      // Drži izdelek v vrteči mizi
              R    "Y3/3_OdpiranjeDržalaKomada"
   END_STEP
   TRANSITION Trans34 FROM ("Odpri klešče", "DRŽI IZDELEK") TO ("VRAČANJE NAZAJ", "Odmik konusa")   // T34
      := "PrijemaloKontaktaOdprto" AND "DrzanjeKontakta";
   END_TRANSITION
   STEP "VRAČANJE NAZAJ":   // S9, max time T#10S, warning time T#7S
      supervision V := (NOT "PrijemaloKontaktaOdprto" OR NOT "SDAT1".oPoz1Dosezena) AND (#"VRAČANJE NAZAJ".T > t#2000MS);
              S    "Y2/1_NalaganjeNazanj"
              R    "Y2/1_NalaganjeNaprej"
              R    "Y1/3_OdmičniCilinderKonusa"
   END_STEP
   TRANSITION Trans41 FROM ("Odmik konusa", "VRAČANJE NAZAJ") TO ("ZAVRTI MIZO", Step36)   // T41
      := ((("FB_KEYENCE_GT2_odmikKonusaKroznika".out >= 57000) AND ("FB_KEYENCE_GT2_ODMIKVARJENJA".out >= 39000)) OR ("AlwaysFALSE" AND "FB_KEYENCE_GT2_ODMIKVARJENJA".oPoz1Dosezena AND "FB_KEYENCE_GT2_odmikKonusaKroznika".oPoz1Dosezena)) AND ("FB_AKD_VrtenjeKroznika".o_BerrStatus = 1);
   END_TRANSITION
   STEP "ZAVRTI MIZO":   // S10, max time T#10S, warning time T#7S
      interlock C := "PozKontaktNazaj" AND "DrzanjeIzmetKontakta" AND "IzmetKontaktaNazaj" AND "PozKontaktNazaj" AND "Y1/4_odmičniCilinderVarjenje_GOR";
      (C)     S    "db_AKD".KROZNIK.PODATKI.ServoGo
   END_STEP
   STEP "ZAKLEP KONUSA":   // S11, max time T#10S, warning time T#7S
              S    "Y1/3_OdmičniCilinderKonusa"
   END_STEP
   STEP "PODAJANJE PLOŠČICE":   // S14, max time T#10S, warning time T#7S
      supervision V := (NOT "SDAT1".oPoz1Dosezena OR NOT "PozKontaktNaKoncuLetve") AND (#"PODAJANJE PLOŠČICE".T > t#2000MS);
              S    "Y2/1_dovajanjePlosciceNazaj"
              R    "Y2_1_dovajanjePlosciceNaprej"
   END_STEP
   TRANSITION Trans38 FROM "PODAJANJE PLOŠČICE" TO "ZAČETEK NOVEGA CIKLA"   // T38: SDAT VREDNOSTI <> 0
      := "SDAT1".oPoz1Dosezena AND "PozKontaktNaKoncuLetve" AND ("SDAT1".out <> 0.0) AND ("SDAT2".out <> 0.0);
   END_TRANSITION
   STEP Step36:   // S36, max time T#10S, warning time T#7S
      interlock C := "PozKontaktNaKoncuLetve" AND "SDAT1".oPoz1Dosezena;
      // Zapri prijemalo
      (C)     R    "Y3/1_PrijemaloKontaktaOdpri"
   END_STEP
   TRANSITION Trans43 FROM ("ZAVRTI MIZO", Step36) TO (Step40, Step37)   // T43
      := NOT "db_AKD".KROZNIK.PODATKI.ServoGo AND "TON_MOTOR".Q AND "DB_PODATKI".KROZNA_MIZA.IzdelekPrisotenArray[5];
   END_TRANSITION
   TRANSITION Trans55 FROM ("ZAVRTI MIZO", Step36) TO "Izdelek ni bil prisoten"   // T55
      := NOT "db_AKD".KROZNIK.PODATKI.ServoGo AND "TON_MOTOR".Q AND NOT "DB_PODATKI".KROZNA_MIZA.IzdelekPrisotenArray[5];
   END_TRANSITION
   STEP "Zakasnitev varjenja":   // S35, max time T#10S, warning time T#7S
      supervision V := ((NOT "EndOfSequency_WC" AND "AlwaysFALSE") OR NOT "FB_KEYENCE_GT2_ODMIKVARJENJA".oPoz4Dosezena) AND (#"Zakasnitev varjenja".T > t#2000MS);
   END_STEP
   TRANSITION Trans19 FROM "Zakasnitev varjenja" TO "Dvig elektrode"   // T19
      := ("EndOfSequency_WC" AND NOT "WeldFault" AND "FB_KEYENCE_GT2_ODMIKVARJENJA".oPoz4Dosezena) OR ("WeldFault" AND "FB_KEYENCE_GT2_ODMIKVARJENJA".oPoz4Dosezena) OR NOT "ExternalWeldOn";
   END_TRANSITION
   STEP "ZAČETEK NOVEGA CIKLA":   // S31, max time T#10S, warning time T#7S
      supervision V := (NOT "PozKontaktNaKoncuLetve" OR NOT "PrisotnostTraka" OR NOT "FB_IOL_IFM_SV_DB".oPretokOK OR NOT "FB_IOL_IFM_SV_DB".oTempOK OR "NapakaCiscenjaElektrode" OR "NapakaOdvijanjaTrau" OR ("FB_TekociTrak_DB".stat_skatla1Polna AND "FB_TekociTrak_DB".stat_skatla2Polna)) AND (#"ZAČETEK NOVEGA CIKLA".T > t#2000MS);
   END_STEP
   TRANSITION Trans48 FROM "ZAČETEK NOVEGA CIKLA" TO Step38   // T48
      := NOT "STEVEC_KONEC_TRAKA_DOSEZEN" AND "FB_IOL_IFM_SV_DB".oPretokOK AND "FB_IOL_IFM_SV_DB".oTempOK AND NOT "NapakaCiscenjaElektrode" AND NOT "NapakaOdvijanjaTrau" AND (NOT "FB_TekociTrak_DB".stat_skatla1Polna OR NOT "FB_TekociTrak_DB".stat_skatla2Polna);
   END_TRANSITION
   STEP Step38:   // S38, max time T#10S, warning time T#7S
      supervision V := NOT "PozKontaktNaKoncuLetve" AND (#Step38.T > t#3000MS);
   END_STEP
   TRANSITION Trans45 FROM Step38 TO Step43   // T45
      := "SDAT1".oPoz1Dosezena AND "PozKontaktNaKoncuLetve" AND NOT "DB_PODATKI".KROZNA_MIZA.IzdelekPrisoten.%X7;
   END_TRANSITION
   TRANSITION Trans47 FROM Step38 TO Step41   // T47: Izdelek prisoten v mizi
      := "DB_PODATKI".KROZNA_MIZA.IzdelekPrisoten.%X7;
   END_TRANSITION
   STEP Step43:   // S43, max time T#10S, warning time T#7S
              R    "DB_VARJENJE".PODATKI.input.ZajtevaZaVarjenje
   END_STEP
   TRANSITION Trans52 FROM Step43 TO ("Odpri Držanje komada", "Zapiranje klešč")   // T52
      := #Step43.T > t#20MS;
   END_TRANSITION
   STEP IZMET:   // S32, max time T#10S, warning time T#7S
              L    "Y4/3_OdpiranjeIzmetaKontakta",T#50mS
              L    "Y5/3_IzmetKomadov", T#50mS
   END_STEP
   TRANSITION Trans46 FROM IZMET TO "NALAGANJE PLOŠČICE/KOMADA"   // T46
      := (#IZMET.T > t#100MS) AND "SDAT1".oPoz1Dosezena;
   END_TRANSITION
   STEP Step41:   // S41, max time T#10S, warning time T#7S
   END_STEP
   TRANSITION Trans49 FROM Step41 TO ("VRAČANJE NAZAJ", "Odmik konusa")   // T49
      := #Step41.T > t#20MS;
   END_TRANSITION
   STEP Step30:   // S30, max time T#10S, warning time T#7S
   END_STEP
   TRANSITION Trans22 FROM Step30 TO "POZ ZAVARJENO"   // T22
      := TRUE;
   END_TRANSITION
   STEP Step37:   // S37, max time T#10S, warning time T#7S
   END_STEP
   TRANSITION Trans37 FROM Step37 TO ("ZAKLEP KONUSA", "IZMET KOSOV", "Poravnava Naprej_1", "Vlaganje ploščice_1", PODAJANJE_1)   // T37: Počakaj da se motor odvrti
      := (#Step37.T > t#20MS) AND ("DB_PODATKI".KROZNA_MIZA.IzdelekPrisoten.%X7 OR "AlwaysTRUE") AND "FB_AKD_DB_RezanjePodajanje".iAKD.PODATKI_TO_SIEMENS.DriveStopen;
   END_TRANSITION
   STEP Step40:   // S40, max time T#10S, warning time T#7S
      supervision V := NOT "PozKontaktNaKoncuLetve" AND (#Step40.T > t#2000MS);
   END_STEP
   TRANSITION Trans44 FROM Step40 TO ("Zapiranje klešč_1", "Odpri Držanje komada_1", "ZAKLEP KONUSA_1")   // T44
      := NOT "DB_PODATKI".KROZNA_MIZA.IzdelekPrisoten.%X7 AND (#Step40.T > t#20MS) AND "PozKontaktNaKoncuLetve";
   END_TRANSITION
   TRANSITION Trans53 FROM Step40 TO "VRAČANJE NAZAJ_1"   // T53
      := "AlwaysTRUE" AND (#Step40.T > t#100MS) AND "DB_PODATKI".KROZNA_MIZA.IzdelekPrisoten.%X7;
   END_TRANSITION
   STEP "Odpri klešče_1":   // S21, max time T#10S, warning time T#7S
      supervision V := NOT "PrijemaloKontaktaOdprto" AND (#"Odpri klešče_1".T > t#2000MS);
              S    "Y3/1_PrijemaloKontaktaOdpri"
              S    "DB_PODATKI".KROZNA_MIZA.IzdelekPrisoten.%X7
   END_STEP
   STEP "Vstavljanje v mizo_1":   // S15, max time T#10S, warning time T#7S
      interlock C := "FB_KEYENCE_GT2_odmikKonusaKroznika".oPoz2Dosezena;
      supervision V := (NOT "PrijemaloKontaktaZaprto" OR NOT "SDAT1".oPoz2Dosezena) AND (#"Vstavljanje v mizo_1".T > t#2000MS);
      (C)     S    "Y2/1_NalaganjeNaprej"
              R    "Y2/1_NalaganjeNazanj"
   END_STEP
   TRANSITION Trans35 FROM "Vstavljanje v mizo_1" TO Step42   // T35
      := "PrijemaloKontaktaZaprto" AND "SDAT1".oPoz2Dosezena;
   END_TRANSITION
   STEP "Zapiranje klešč_1":   // S6, max time T#10S, warning time T#7S
      interlock C := "PozKontaktNaKoncuLetve";
      (C)     R    "Y3/1_PrijemaloKontaktaOdpri"
   END_STEP
   STEP "Odpri Držanje komada_1":   // S13, max time T#10S, warning time T#7S
      supervision V := "DrzanjeKontakta" AND (#"Odpri Držanje komada_1".T > t#2000MS);
      // OdpriDržanjeKomada -
              S    "Y3/3_OdpiranjeDržalaKomada"
   END_STEP
   STEP "DRŽI IZDELEK_1":   // S33, max time T#10S, warning time T#7S
      supervision V := NOT "DrzanjeKontakta" AND (#"DRŽI IZDELEK_1".T > t#2000MS);
      // Drži izdelek v vrteči mizi
              R    "Y3/3_OdpiranjeDržalaKomada"
   END_STEP
   TRANSITION Trans40 FROM ("Odpri klešče_1", "DRŽI IZDELEK_1") TO "VRAČANJE NAZAJ_1"   // T40
      := "PrijemaloKontaktaOdprto" AND "DrzanjeKontakta";
   END_TRANSITION
   STEP "VRAČANJE NAZAJ_1":   // S34, max time T#10S, warning time T#7S
      supervision V := (NOT "PrijemaloKontaktaOdprto" OR NOT "SDAT1".oPoz1Dosezena) AND (#"VRAČANJE NAZAJ_1".T > t#2000MS);
              S    "Y2/1_NalaganjeNazanj"
              R    "Y2/1_NalaganjeNaprej"
   END_STEP
   STEP "ZAKLEP KONUSA_1":   // S39, max time T#10S, warning time T#7S
              S    "Y1/3_OdmičniCilinderKonusa"
   END_STEP
   TRANSITION Trans33 FROM ("Zapiranje klešč_1", "Odpri Držanje komada_1", "ZAKLEP KONUSA_1") TO "Vstavljanje v mizo_1"   // T33: Prijemalo zaprto
      := "PrijemaloKontaktaZaprto" AND NOT "DrzanjeKontakta" AND "ZaporaIzdelka";
   END_TRANSITION
   STEP Step42:   // S42, max time T#10S, warning time T#7S
              S    "Y3/1_PrijemaloKontaktaOdpri"
              S    "DB_PODATKI".KROZNA_MIZA.IzdelekPrisoten.%X7
   END_STEP
   TRANSITION Trans54 FROM Step42 TO ("DRŽI IZDELEK_1", "Odpri klešče_1")   // T54
      := TRUE;
   END_TRANSITION
   STEP "Izdelek ni bil prisoten":   // S44, max time T#10S, warning time T#7S
   END_STEP
   TRANSITION Trans56 FROM "Izdelek ni bil prisoten" TO "ZAČETEK NOVEGA CIKLA"   // T56, jump
      := TRUE;
   END_TRANSITION
   STEP "Poravnava Naprej_1":   // S46, max time T#10S, warning time T#7S
              S    "Y2/3_PozicioniranjeKontaktovNaprej"
              R    "Y2/3_PozicioniranjeKontaktovNazaj"
              S    "1Y1_OdklepZapore"
   END_STEP
   STEP "Vlaganje ploščice_1":   // S48, max time T#10S, warning time T#7S
      interlock C := "FB_KEYENCE_GT2_ODMIKVARJENJA".oPoz1Dosezena;
      supervision V := NOT "SDAT2".oPoz2Dosezena AND (#"Vlaganje ploščice_1".U > t#2000MS);
              S    "Y2_1_dovajanjePlosciceNaprej"
              R    "Y2/1_dovajanjePlosciceNazaj"
   END_STEP
   STEP "ZVAR NOK":   // S50, max time T#10S, warning time T#7S
      supervision V := "IEC_Counter_0_DB_1".QU;
              R    "DB_PODATKI".KROZNA_MIZA.IzdelekZavarjen.%X5
              N    "DB_PODATKI".KROZNA_MIZA.StatusIzdelkaVarjenje[5] := 1
              S    "DB_HMI".Varjenje.ResetWithWC
   END_STEP
   TRANSITION Trans59 FROM "ZVAR NOK" TO "Zakasnitev varjenja"   // T59
      := NOT "IEC_Counter_0_DB_1".QU;
   END_TRANSITION
   STEP "Zvar  OK":   // S51, max time T#10S, warning time T#7S
              S    "DB_PODATKI".KROZNA_MIZA.IzdelekZavarjen.%X5
              N    "DB_PODATKI".KROZNA_MIZA.StatusIzdelkaVarjenje[5] := 10
   END_STEP
   TRANSITION Trans60 FROM "Zvar  OK" TO "Zakasnitev varjenja"   // T60
      := TRUE;
   END_TRANSITION
   STEP Step52:   // S52, max time T#10S, warning time T#7S
   END_STEP
   TRANSITION Trans62 FROM Step52 TO (Step45, REZANJE)   // T62
      := TRUE;
   END_TRANSITION
   STEP Step16:   // S16, max time T#10S, warning time T#7S
      supervision V := NOT "EndOfSequency_WC" AND (#Step16.T > t#1000MS);
   END_STEP
   TRANSITION Trans50 FROM Step16 TO "Zvar  OK"   // T50
      := "EndOfSequency_WC" AND NOT "WeldFault";
   END_TRANSITION
   TRANSITION Trans58 FROM Step16 TO "ZVAR NOK"   // T58
      := "WeldFault";
   END_TRANSITION
   STEP Step54:   // S54, max time T#10S, warning time T#7S
      // Ploščica Odrezana - setiraj bit
              N    "db_AKD".REZANJEPODAJANJE.PODATKI.PloscicaOdrezana := True
   END_STEP
   TRANSITION Trans64 FROM Step54 TO END   // T64
      := TRUE;
   END_TRANSITION
   STEP "RESET VSEGA":   // S2, max time T#10S, warning time T#7S
      // RESET ENOTE
              R    "Y2/1_NalaganjeNaprej"
              R    "Y2/1_NalaganjeNazanj"
              S    "Y3/1_PrijemaloKontaktaOdpri"
              R    "Y2/3_PozicioniranjeKontaktovNazaj"
              S    "Y1/3_OdmičniCilinderKonusa"
              R    "Y3/3_OdpiranjeDržalaKomada"
              R    "Y4/3_OdpiranjeIzmetaKontakta"
              R    "Y5/3_IzmetKomadov"
              S    "Y1/4_odmičniCilinderVarjenje_GOR"
              S    "1Y1_OdklepZapore"
              S    "Y2/1_dovajanjePlosciceNazaj"
              R    "Y2_1_dovajanjePlosciceNaprej"
              R    "db_AKD".REZANJEPODAJANJE.PODATKI.Odrezano
              R    "db_AKD".REZANJEPODAJANJE.PODATKI.Podano
              R    "Y2/1_dovajanjePlosciceNazaj"
              R    "Y2_1_dovajanjePlosciceNaprej"
              R    "Y2/3_PozicioniranjeKontaktovNaprej"
              S    "Y2/3_PozicioniranjeKontaktovNazaj"
              R    "Y2_1_dovajanjePlosciceNaprej"
              R    "Y2/1_dovajanjePlosciceNazaj"
              R    "db_AKD".REZANJEPODAJANJE.PODATKI.Odrezano
              R    "db_AKD".REZANJEPODAJANJE.PODATKI.Podano
              R    "db_AKD".REZANJEPODAJANJE.PODATKI.ZahtevaPoPodajanju
              R    "db_AKD".REZANJEPODAJANJE.PODATKI.ZahtevaPoRezanju
              R    "DB_VARJENJE".PODATKI.input.ZajtevaZaVarjenje
              R    "Y1/4_odmičniCilinderVarjenjeDOL"
              S    "Y3/1_PrijemaloKontaktaOdpri"
              R    "DB_VARJENJE".PODATKI.input.ZajtevaZaVarjenje
              R    "DB_HMI".Varjenje.ResetWithWC
              R    "Y5/3_IzmetKomadov"
   END_STEP
   TRANSITION Trans28 FROM "RESET VSEGA" TO IZMET   // T28: OK
      := TRUE;
   END_TRANSITION
   STEP "Odmik vilic":   // S27, max time T#10S, warning time T#7S
      supervision V := (NOT "SDAT2".oPoz1Dosezena OR (NOT "TimerReady" AND "AlwaysFALSE") OR ("WeldFault" AND "AlwaysFALSE") OR NOT "SpotSelectionTakeOver") AND (#"Odmik vilic".T > t#2000MS);
              S    "Y2/1_dovajanjePlosciceNazaj"
              R    "Y2_1_dovajanjePlosciceNaprej"
              N    "db_AKD".REZANJEPODAJANJE.PODATKI.PloscicaOdrezana := false
   END_STEP
   TRANSITION Trans26 FROM ("VRAČANJE NAZAJ_1", "Poravnava nazaj", "Odmik vilic") TO (Varjenje, Step52)   // T26: Vilice v izhodišču + pdoajanje v izhodišču
      := ("SDAT2".oPoz1Dosezena OR ("SDAT2".out <= 60.0)) AND "PozKontaktNazaj" AND (("TimerReady" AND NOT "WeldFault") OR "AlwaysTRUE") AND "SpotSelectionTakeOver" AND "FB_KEYENCE_GT2_ODMIKVARJENJA".oPoz3Dosezena AND ("SDAT1".oPoz1Dosezena OR ("SDAT1".out <= 50.0) OR "AlwaysTRUE") AND "FB_KEYENCE_GT2_odmikKonusaKroznika".oPoz2Dosezena AND ("FB_AKD_DB_RezanjePodajanje".o_BerrStatus = 1);
   END_TRANSITION
   STEP "Odmik konusa":   // S22, max time T#10S, warning time T#7S
              R    "Y1/3_OdmičniCilinderKonusa"
   END_STEP
   STEP PODAJANJE_1:   // S47, max time T#10S, warning time T#7S
              S    "db_AKD".REZANJEPODAJANJE.PODATKI.Podano
              L    "db_AKD".REZANJEPODAJANJE.PODATKI.ZahtevaPoPodajanju, T#50mS
   END_STEP
   TRANSITION Trans36 FROM PODAJANJE_1 TO Step53   // T36
      := NOT "FB_AKD_DB_RezanjePodajanje".bServoGo AND "TON_REZANJEPODAJANJE".Q AND NOT "db_AKD".REZANJEPODAJANJE.PODATKI.vPODAJANJU AND (#PODAJANJE_1.T > t#10MS);
   END_TRANSITION
   STEP Step53:   // S53, max time T#10S, warning time T#7S
   END_STEP
   TRANSITION Trans24 FROM ("IZMET KOSOV", "ZAKLEP KONUSA", "Poravnava Naprej_1", "Vlaganje ploščice_1", Step53) TO "Spust Elektrode"   // T24: Izmet Nazaj in KONUS zaklenjen
      := "DrzanjeIzmetKontakta" AND "IzmetKontaktaNazaj" AND "FB_KEYENCE_GT2_odmikKonusaKroznika".oPoz2Dosezena AND "PozKontaktNaprej" AND "SDAT2".oPoz2Dosezena AND (#"IZMET KOSOV".T > t#50MS);
   END_TRANSITION
   STEP Step49:   // S49, max time T#10S, warning time T#7S
              S    "Y2_1_dovajanjePlosciceNaprej"
              R    "Y2/1_dovajanjePlosciceNazaj"
   END_STEP
   TRANSITION Trans51 FROM Step49 TO "Izdelek ni bil prisoten"   // T51
      := TRUE;
   END_TRANSITION

   // permanent post-instructions
   NETWORK 1
   TITLE = ODKLENI LIN PROGO
      "1Y1_OdklepZapore" := ("SDAT1".out >= 19.5) OR (("SDAT1".out < 19.5) AND NOT "PozKontaktNaKoncuLetve");
   NETWORK 2
   TITLE = VSTAVLJANJE KOSA V MIZO
   NETWORK 3
      IF "AlwaysFALSE" THEN
          "FB_Alarms_DB_1"(I_FAULT_RESET := "ResetNapake",   // "FB_Alarms"
                           I_Alarm_0 := "FB_GL_PROGRAM_DB"."Spust Elektrode".X AND NOT "FB_KEYENCE_GT2_ODMIKVARJENJA".bBDC3,
                           I_Alarm_1 := ("FB_FESTO_SDE1_DB".oPritisk < 6.0) AND "AlwaysFALSE",
                           I_Alarm_2 := NOT "PrisotnostTraka" AND "AlwaysFALSE",
                           I_Alarm_3 := #"Vstavljanje v mizo_1".VA,
                           I_Alarm_4 := #"Vstavljanje v mizo_1".VS,
                           I_Alarm_5 := #"Vstavljanje v mizo_1".V0,
                           I_Alarm_6 := #"Vstavljanje v mizo_1".LA,
                           I_Alarm_7 := #"Vstavljanje v mizo_1".S1);
      END_IF;
   NETWORK 4
   TITLE = ŠTEVEC
      "STEVECKOSOV_PO_KONCU_TRAKU".CTU(CU := NOT "PrisotnostTraka" AND #"IZMET KOSOV".X,
                              R := "PrisotnostTraka",
                              PV := 110);
      "STEVEC_KONEC_TRAKA_DOSEZEN" := "STEVECKOSOV_PO_KONCU_TRAKU".Q;
      IF NOT "PrisotnostTraka" AND NOT "STEVEC_KONEC_TRAKA_DOSEZEN" THEN "StatusPrisotnostiTraku" := 10; END_IF;
      IF NOT "PrisotnostTraka" AND "STEVEC_KONEC_TRAKA_DOSEZEN" THEN "StatusPrisotnostiTraku" := 0; END_IF;
      IF "PrisotnostTraka" THEN "StatusPrisotnostiTraku" := 1; END_IF;
   NETWORK 5
   TITLE = Odvijanje traku
      "MotorOdvijanjeTraku" := "SenzorStartOdvijanje";
   NETWORK 6
   TITLE = ŠTEVCI - števec zavarjen 10, error 11
      #_w1 := #"IZMET KOSOV".X AND NOT "DB_PODATKI".KROZNA_MIZA.MerkerjiKoraka[0];   // rising edge of #"IZMET KOSOV".X
      "DB_PODATKI".KROZNA_MIZA.MerkerjiKoraka[0] := #"IZMET KOSOV".X;
      #_w2 := #_w1 AND ("DB_PODATKI".KROZNA_MIZA.StatusIzdelkaVarjenje[1] = 10) AND "DB_PODATKI".KROZNA_MIZA.IzdelekPrisoten.%X1;
      IF #_w2 THEN
          "DB_STEVCI"."STEVCI VARJENJE".SKUPAJOK := "DB_STEVCI"."STEVCI VARJENJE".SKUPAJOK + 1;
          "DB_STEVCI"."STEVCI VARJENJE".ZavarjenoOK := "DB_STEVCI"."STEVCI VARJENJE".ZavarjenoOK + 1;
      END_IF;
      #onemogoci := #_w2;
      IF #_w2 AND NOT "PolnjenjeSkatle1" THEN
          "DB_STEVCI".STEVEC_SKATEL.SKATLA1 := "DB_STEVCI".STEVEC_SKATEL.SKATLA1 + 1;
      END_IF;
      IF #_w2 AND "PolnjenjeSkatle1" THEN
          "DB_STEVCI".STEVEC_SKATEL.SKATLA2 := "DB_STEVCI".STEVEC_SKATEL.SKATLA2 + 1;
      END_IF;
      IF #_w1 AND NOT #onemogoci AND ("DB_PODATKI".KROZNA_MIZA.IzdelekZavarjen <> 10) AND "DB_PODATKI".KROZNA_MIZA.IzdelekPrisoten.%X1 THEN
          "DB_STEVCI"."STEVCI VARJENJE".ZavarjenoNOK := "DB_STEVCI"."STEVCI VARJENJE".ZavarjenoNOK + 1;
          "DB_STEVCI".STEVEC_SKATEL.SKATLA_SLABI := "DB_STEVCI".STEVEC_SKATEL.SKATLA_SLABI + 1;
          "DB_STEVCI"."STEVCI VARJENJE".SKUPAJNOK := "DB_STEVCI"."STEVCI VARJENJE".SKUPAJNOK + 1;
      END_IF;
END_FUNCTION_BLOCK

FUNCTION_BLOCK "FB_AKD"   // FB6, LAD
{ S7_Optimized_Access := 'TRUE' }
VERSION : 0.1
   VAR_INPUT
      bServoEnable : Bool;
      iNastavitevHitrosti : Int;
      dNastavitevPozicije : DInt;
      bPogojiZaVKLOP : Bool;
      iAKD : "AKD_TO_SIEMENS";
      ResetNapake : Bool;
      iStPrograma : Word;
   END_VAR
   VAR_OUTPUT
      oAKD : "SIEMENS_TO_AKD";
      AKDcurrPos : DInt;
      o_BerrStatus : Byte;
      rAKDpos : Real;
   END_VAR
   VAR_IN_OUT
      iStartHoming : Bool;
      bServoGo : Bool;
   END_VAR
   VAR
      TIMER_ON : Array[0..4] of TON_TIME;
      diHitrost : Real;
      dwHitrostRez : Real;
      ServoHommed : Bool;
   END_VAR
   VAR RETAIN
      merker : Array[0..1] of Bool;
   END_VAR
   VAR
      OmogociHome : Bool;
   END_VAR
   VAR_TEMP   // added for the SCL form of the ladder/FBD networks
      _w1 : Bool;
   END_VAR
BEGIN

REGION Network 1: Bool
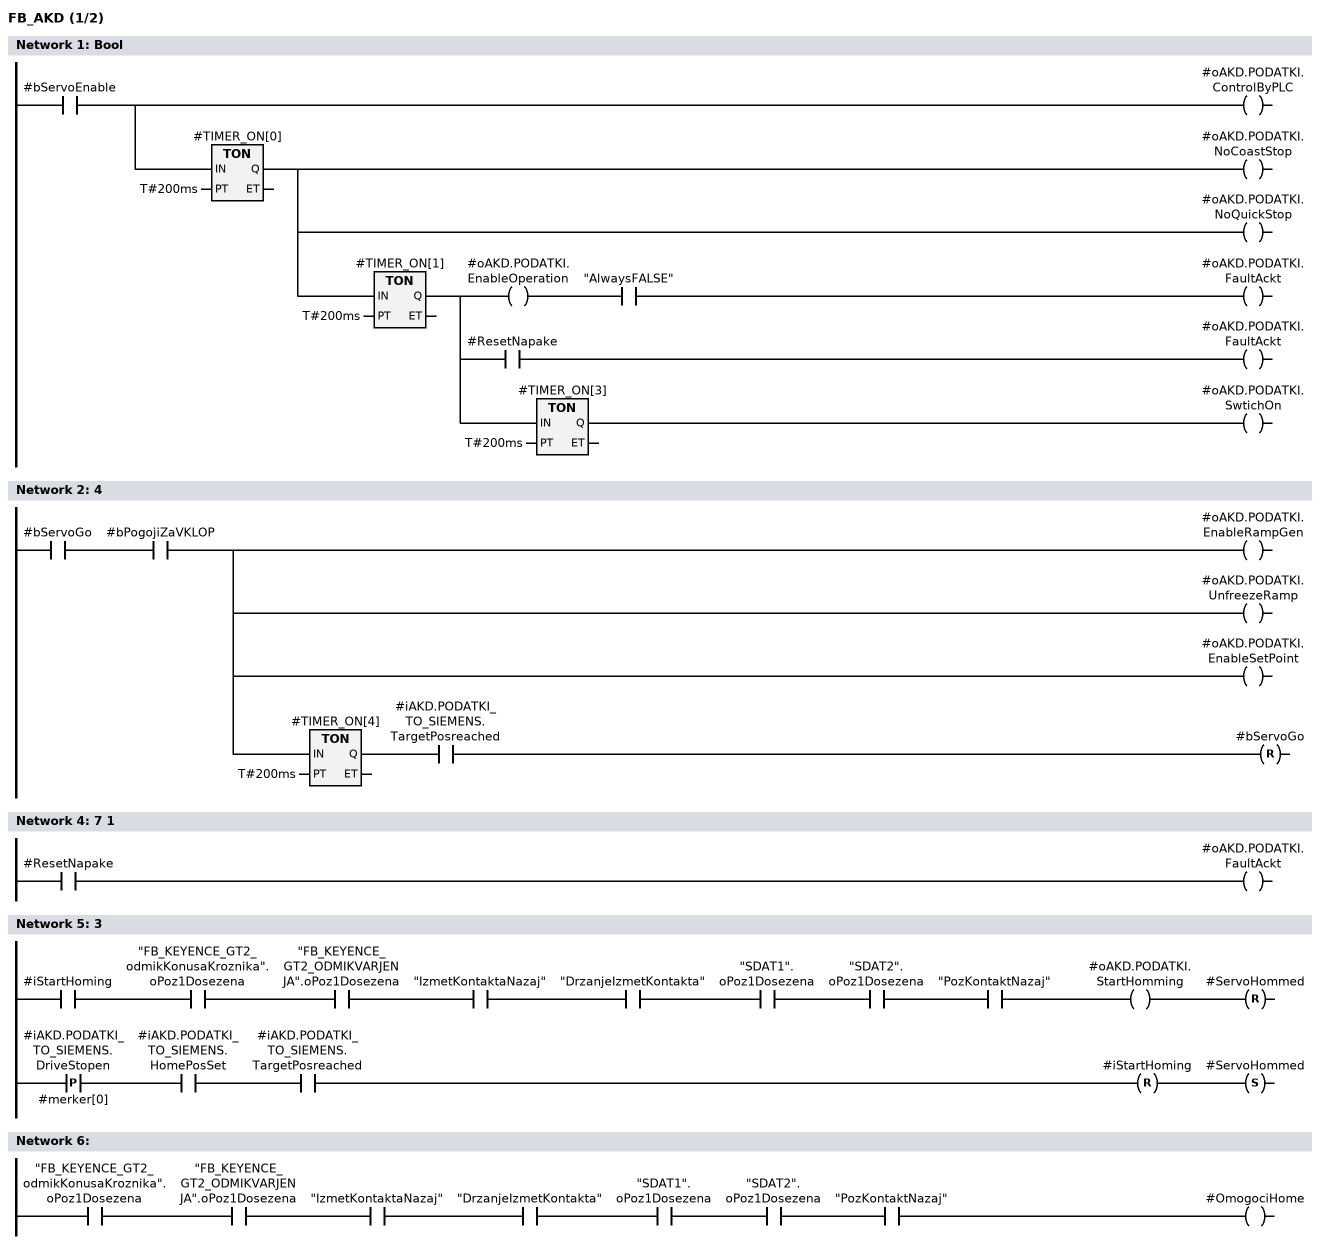
   #oAKD.PODATKI.ControlByPLC := #bServoEnable;
   #TIMER_ON[0].TON(IN := #bServoEnable, PT := T#200ms);
   #oAKD.PODATKI.NoCoastStop := #TIMER_ON[0].Q;
   #oAKD.PODATKI.NoQuickStop := #TIMER_ON[0].Q;
   #TIMER_ON[1].TON(IN := #TIMER_ON[0].Q, PT := T#200ms);
   #oAKD.PODATKI.EnableOperation := #TIMER_ON[1].Q;
   #oAKD.PODATKI.FaultAckt := #TIMER_ON[1].Q AND "AlwaysFALSE";
   #oAKD.PODATKI.FaultAckt := #TIMER_ON[1].Q AND #ResetNapake;
   #TIMER_ON[3].TON(IN := #TIMER_ON[1].Q, PT := T#200ms);
   #oAKD.PODATKI.SwtichOn := #TIMER_ON[3].Q;
END_REGION

REGION Network 2: 4
   #oAKD.PODATKI.EnableRampGen := #bServoGo AND #bPogojiZaVKLOP;
   #oAKD.PODATKI.UnfreezeRamp := #oAKD.PODATKI.EnableRampGen;
   #oAKD.PODATKI.EnableSetPoint := #oAKD.PODATKI.EnableRampGen;
   #TIMER_ON[4].TON(IN := #oAKD.PODATKI.EnableRampGen, PT := T#200ms);
   IF #TIMER_ON[4].Q AND #iAKD.PODATKI_TO_SIEMENS.TargetPosreached THEN #bServoGo := FALSE; END_IF;
END_REGION

REGION Network 3 (SCL)
   //PretvorbaHitrosti
   #diHitrost := INT_TO_REAL(#iNastavitevHitrosti);
   #dwHitrostRez :=((#diHitrost * 4294967295/12000));
   #oAKD.PODATKI.MDI_VELOCITY := REAL_TO_DINT(#dwHitrostRez); //hitrost


   // Operation mode
   #oAKD.PODATKI.MDI_MOD := 16#00_00; //0 - relativni 1//aboslutni gib
   #oAKD.PODATKI.SATANW := #iStPrograma;   //OutputTask

   //pretvorba poziij
   #AKDcurrPos := (#iAKD.PODATKI_TO_SIEMENS.ActualPos * 5 )/ 65536;
   #rAKDpos:= (#iAKD.PODATKI_TO_SIEMENS.ActualPos) / 65536.00;
   //nastavljanjePozicije
   //nastavljanje pozicije
   #oAKD.PODATKI.MDI_TARPOS := (65536 * #dNastavitevPozicije / 5);
END_REGION

REGION Network 4: 7 1
   RUNG wire#powerrail
      Contact( #ResetNapake )
      Coil( #oAKD.PODATKI.FaultAckt )
   END_RUNG
   // the same network as SCL:
   #oAKD.PODATKI.FaultAckt := #ResetNapake;
END_REGION

REGION Network 5: 3
   RUNG wire#powerrail
      Contact( #iStartHoming )
      Contact( "FB_KEYENCE_GT2_odmikKonusaKroznika".oPoz1Dosezena )
      Contact( "FB_KEYENCE_GT2_ODMIKVARJENJA".oPoz1Dosezena )
      Contact( "IzmetKontaktaNazaj" )
      Contact( "DrzanjeIzmetKontakta" )
      Contact( "SDAT1".oPoz1Dosezena )
      Contact( "SDAT2".oPoz1Dosezena )
      Contact( "PozKontaktNazaj" )
      Coil( #oAKD.PODATKI.StartHomming )
      R_Coil( #ServoHommed )
   END_RUNG
   RUNG wire#powerrail
      P_Contact(operand := #iAKD.PODATKI_TO_SIEMENS.DriveStopen, bit := #merker[0])
      Contact( #iAKD.PODATKI_TO_SIEMENS.HomePosSet )
      Contact( #iAKD.PODATKI_TO_SIEMENS.TargetPosreached )
      R_Coil( #iStartHoming )
      S_Coil( #ServoHommed )
   END_RUNG
   // the same network as SCL:
   #oAKD.PODATKI.StartHomming := #iStartHoming AND "FB_KEYENCE_GT2_odmikKonusaKroznika".oPoz1Dosezena AND "FB_KEYENCE_GT2_ODMIKVARJENJA".oPoz1Dosezena AND "IzmetKontaktaNazaj" AND "DrzanjeIzmetKontakta" AND "SDAT1".oPoz1Dosezena AND "SDAT2".oPoz1Dosezena AND "PozKontaktNazaj";
   IF #oAKD.PODATKI.StartHomming THEN #ServoHommed := FALSE; END_IF;
   #_w1 := #iAKD.PODATKI_TO_SIEMENS.DriveStopen AND NOT #merker[0];   // rising edge of #iAKD.PODATKI_TO_SIEMENS.DriveStopen
   #merker[0] := #iAKD.PODATKI_TO_SIEMENS.DriveStopen;
   IF #_w1 AND #iAKD.PODATKI_TO_SIEMENS.HomePosSet AND #iAKD.PODATKI_TO_SIEMENS.TargetPosreached THEN
       #iStartHoming := FALSE;
       #ServoHommed := TRUE;
   END_IF;
END_REGION

REGION Network 6
   RUNG wire#powerrail
      Contact( "FB_KEYENCE_GT2_odmikKonusaKroznika".oPoz1Dosezena )
      Contact( "FB_KEYENCE_GT2_ODMIKVARJENJA".oPoz1Dosezena )
      Contact( "IzmetKontaktaNazaj" )
      Contact( "DrzanjeIzmetKontakta" )
      Contact( "SDAT1".oPoz1Dosezena )
      Contact( "SDAT2".oPoz1Dosezena )
      Contact( "PozKontaktNazaj" )
      Coil( #OmogociHome )
   END_RUNG
   // the same network as SCL:
   #OmogociHome := "FB_KEYENCE_GT2_odmikKonusaKroznika".oPoz1Dosezena AND "FB_KEYENCE_GT2_ODMIKVARJENJA".oPoz1Dosezena AND "IzmetKontaktaNazaj" AND "DrzanjeIzmetKontakta" AND "SDAT1".oPoz1Dosezena AND "SDAT2".oPoz1Dosezena AND "PozKontaktNazaj";
END_REGION

REGION Network 7: ERROR STATUS
END_REGION

REGION Network 8
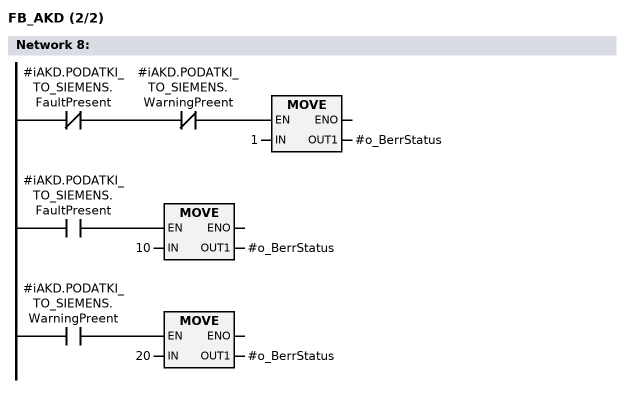
   RUNG wire#powerrail
      I_Contact( #iAKD.PODATKI_TO_SIEMENS.FaultPresent )
      I_Contact( #iAKD.PODATKI_TO_SIEMENS.WarningPreent )
      Move(in := 1, out1 => #o_BerrStatus)
   END_RUNG
   RUNG wire#powerrail
      Contact( #iAKD.PODATKI_TO_SIEMENS.FaultPresent )
      Move(in := 10, out1 => #o_BerrStatus)
   END_RUNG
   RUNG wire#powerrail
      Contact( #iAKD.PODATKI_TO_SIEMENS.WarningPreent )
      Move(in := 20, out1 => #o_BerrStatus)
   END_RUNG
   // the same network as SCL:
   IF NOT #iAKD.PODATKI_TO_SIEMENS.FaultPresent AND NOT #iAKD.PODATKI_TO_SIEMENS.WarningPreent THEN
       #o_BerrStatus := 1;
   END_IF;
   IF #iAKD.PODATKI_TO_SIEMENS.FaultPresent THEN #o_BerrStatus := 10; END_IF;
   IF #iAKD.PODATKI_TO_SIEMENS.WarningPreent THEN #o_BerrStatus := 20; END_IF;
END_REGION
END_FUNCTION_BLOCK

FUNCTION_BLOCK "FB_STARTUP"   // FB7, LAD
{ S7_Optimized_Access := 'TRUE' }
VERSION : 0.1
   VAR_INPUT
      bHMILifeBit : Bool;
      bHMI_StartUp : Bool;
      icurrHMINb : Int;
   END_VAR
   VAR
      korak : UInt;
      IEC_Timer_0_Instance : TON_TIME;
      IEC_Timer_0_Instance_1 : TON_TIME;
      trenutniKorak : Array[0..100] of Bool;
   END_VAR
   VAR RETAIN
      merkers : Array[0..100] of Bool;
      T_ON : Array[0..100] of TON_TIME;
   END_VAR
   VAR
      DeviceState : Struct
         myLADDR : Hw_IoSystem := 260;
         myMODE : UInt := 4;
         returnValue : Int;
         mySTATE : Array[0..1023] of Bool;
      END_STRUCT;
   END_VAR
   VAR_TEMP   // added for the SCL form of the ladder/FBD networks
      _w1 : Bool;
      _w2 : Bool;
   END_VAR
   // // DeviceState.mySTATE[0] : ProfinetIO master
   // // DeviceState.mySTATE[1] : MVK1
   // // DeviceState.mySTATE[2] : MVK2
   // // DeviceState.mySTATE[3] : MVK3
   // // DeviceState.mySTATE[4] : BOSH varilnik
   // // DeviceState.mySTATE[5] : AKD cilinder
   // // DeviceState.mySTATE[6] : Keyence PN-1
   // // DeviceState.mySTATE[7] : AKD vrtljiva miza
   // // DeviceState.mySTATE[8] : AKD elektroda
BEGIN

REGION Network 1
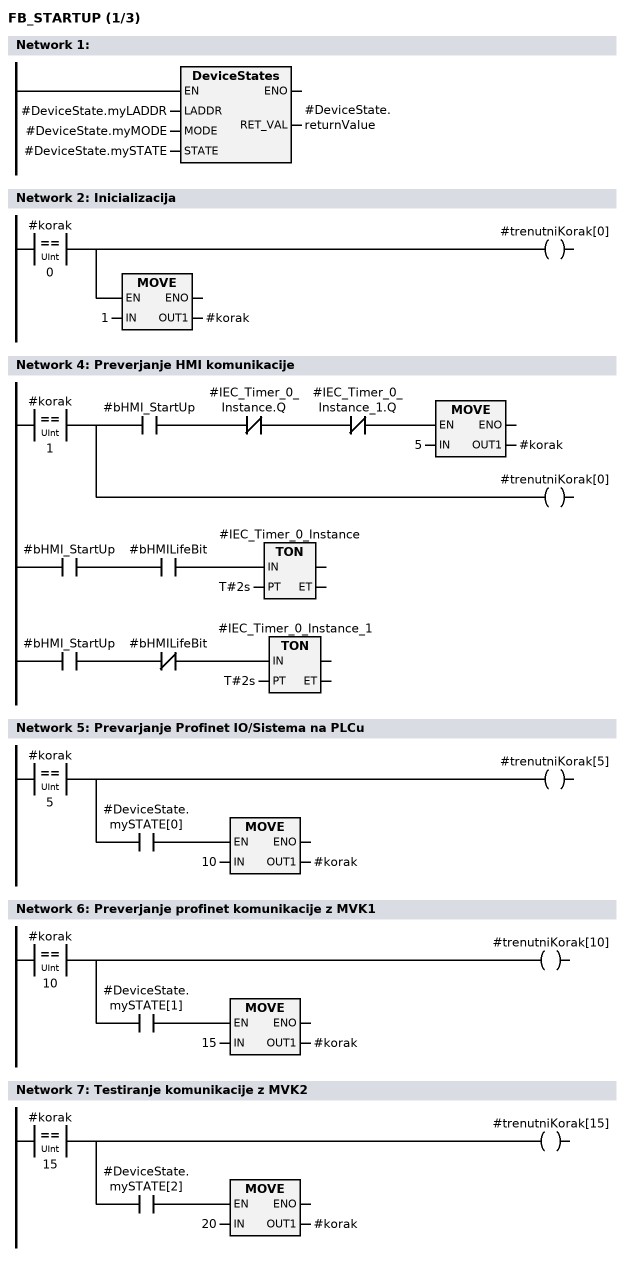
   // no SCL statement known for DeviceStates: written as a call
   #DeviceState.returnValue := DeviceStates(LADDR := #DeviceState.myLADDR,
                           MODE := #DeviceState.myMODE,
                           STATE := #DeviceState.mySTATE);
END_REGION

REGION Network 2: Inicializacija
   RUNG wire#powerrail
      { S7_Templates := "SrcType := UInt" } EQ_Contact(in1 := #korak, in2 := 0)
      wire#w1
      Coil( #trenutniKorak[0] )
   END_RUNG
   RUNG wire#w1
      Move(in := 1, out1 => #korak)
   END_RUNG
   // the same network as SCL:
   #trenutniKorak[0] := #korak = 0;
   IF #korak = 0 THEN #korak := 1; END_IF;
END_REGION

REGION Network 4: Preverjanje HMI komunikacije
   #_w1 := #korak = 1;
   IF #_w1 AND #bHMI_StartUp AND NOT #IEC_Timer_0_Instance.Q AND NOT #IEC_Timer_0_Instance_1.Q THEN
       #korak := 5;
   END_IF;
   #trenutniKorak[0] := #_w1;
   #IEC_Timer_0_Instance(IN := #bHMI_StartUp AND #bHMILifeBit, PT := T#2s);   // TON
   #IEC_Timer_0_Instance_1(IN := #bHMI_StartUp AND NOT #bHMILifeBit, PT := T#2s);   // TON
END_REGION

REGION Network 5: Prevarjanje Profinet IO/Sistema na PLCu
   RUNG wire#powerrail
      { S7_Templates := "SrcType := UInt" } EQ_Contact(in1 := #korak, in2 := 5)
      wire#w1
      Coil( #trenutniKorak[5] )
   END_RUNG
   RUNG wire#w1
      Contact( #DeviceState.mySTATE[0] )
      Move(in := 10, out1 => #korak)
   END_RUNG
   // the same network as SCL:
   #trenutniKorak[5] := #korak = 5;
   IF (#korak = 5) AND #DeviceState.mySTATE[0] THEN #korak := 10; END_IF;
END_REGION

REGION Network 6: Preverjanje profinet komunikacije z MVK1
   RUNG wire#powerrail
      { S7_Templates := "SrcType := UInt" } EQ_Contact(in1 := #korak, in2 := 10)
      wire#w1
      Coil( #trenutniKorak[10] )
   END_RUNG
   RUNG wire#w1
      Contact( #DeviceState.mySTATE[1] )
      Move(in := 15, out1 => #korak)
   END_RUNG
   // the same network as SCL:
   #trenutniKorak[10] := #korak = 10;
   IF (#korak = 10) AND #DeviceState.mySTATE[1] THEN #korak := 15; END_IF;
END_REGION

REGION Network 7: Testiranje komunikacije z MVK2
   RUNG wire#powerrail
      { S7_Templates := "SrcType := UInt" } EQ_Contact(in1 := #korak, in2 := 15)
      wire#w1
      Coil( #trenutniKorak[15] )
   END_RUNG
   RUNG wire#w1
      Contact( #DeviceState.mySTATE[2] )
      Move(in := 20, out1 => #korak)
   END_RUNG
   // the same network as SCL:
   #trenutniKorak[15] := #korak = 15;
   IF (#korak = 15) AND #DeviceState.mySTATE[2] THEN #korak := 20; END_IF;
END_REGION

REGION Network 8: Testiranje komunikacije z MVK3
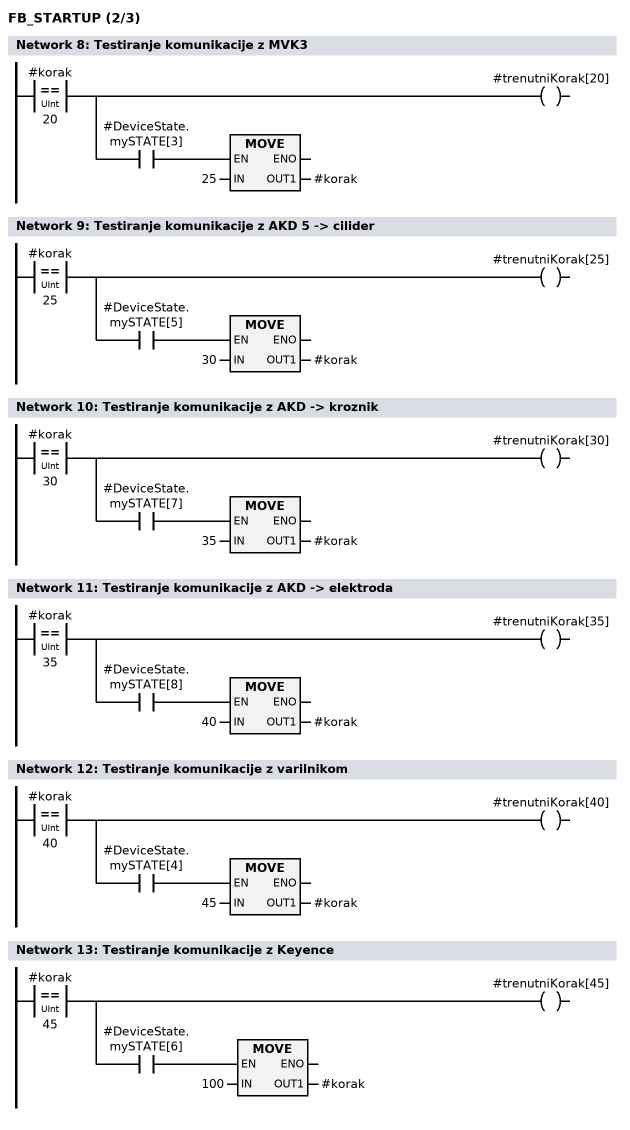
   RUNG wire#powerrail
      { S7_Templates := "SrcType := UInt" } EQ_Contact(in1 := #korak, in2 := 20)
      wire#w1
      Coil( #trenutniKorak[20] )
   END_RUNG
   RUNG wire#w1
      Contact( #DeviceState.mySTATE[3] )
      Move(in := 25, out1 => #korak)
   END_RUNG
   // the same network as SCL:
   #trenutniKorak[20] := #korak = 20;
   IF (#korak = 20) AND #DeviceState.mySTATE[3] THEN #korak := 25; END_IF;
END_REGION

REGION Network 9: Testiranje komunikacije z AKD 5 -> cilider
   RUNG wire#powerrail
      { S7_Templates := "SrcType := UInt" } EQ_Contact(in1 := #korak, in2 := 25)
      wire#w1
      Coil( #trenutniKorak[25] )
   END_RUNG
   RUNG wire#w1
      Contact( #DeviceState.mySTATE[5] )
      Move(in := 30, out1 => #korak)
   END_RUNG
   // the same network as SCL:
   #trenutniKorak[25] := #korak = 25;
   IF (#korak = 25) AND #DeviceState.mySTATE[5] THEN #korak := 30; END_IF;
END_REGION

REGION Network 10: Testiranje komunikacije z AKD -> kroznik
   RUNG wire#powerrail
      { S7_Templates := "SrcType := UInt" } EQ_Contact(in1 := #korak, in2 := 30)
      wire#w1
      Coil( #trenutniKorak[30] )
   END_RUNG
   RUNG wire#w1
      Contact( #DeviceState.mySTATE[7] )
      Move(in := 35, out1 => #korak)
   END_RUNG
   // the same network as SCL:
   #trenutniKorak[30] := #korak = 30;
   IF (#korak = 30) AND #DeviceState.mySTATE[7] THEN #korak := 35; END_IF;
END_REGION

REGION Network 11: Testiranje komunikacije z AKD -> elektroda
   RUNG wire#powerrail
      { S7_Templates := "SrcType := UInt" } EQ_Contact(in1 := #korak, in2 := 35)
      wire#w1
      Coil( #trenutniKorak[35] )
   END_RUNG
   RUNG wire#w1
      Contact( #DeviceState.mySTATE[8] )
      Move(in := 40, out1 => #korak)
   END_RUNG
   // the same network as SCL:
   #trenutniKorak[35] := #korak = 35;
   IF (#korak = 35) AND #DeviceState.mySTATE[8] THEN #korak := 40; END_IF;
END_REGION

REGION Network 12: Testiranje komunikacije z varilnikom
   RUNG wire#powerrail
      { S7_Templates := "SrcType := UInt" } EQ_Contact(in1 := #korak, in2 := 40)
      wire#w1
      Coil( #trenutniKorak[40] )
   END_RUNG
   RUNG wire#w1
      Contact( #DeviceState.mySTATE[4] )
      Move(in := 45, out1 => #korak)
   END_RUNG
   // the same network as SCL:
   #trenutniKorak[40] := #korak = 40;
   IF (#korak = 40) AND #DeviceState.mySTATE[4] THEN #korak := 45; END_IF;
END_REGION

REGION Network 13: Testiranje komunikacije z Keyence
   RUNG wire#powerrail
      { S7_Templates := "SrcType := UInt" } EQ_Contact(in1 := #korak, in2 := 45)
      wire#w1
      Coil( #trenutniKorak[45] )
   END_RUNG
   RUNG wire#w1
      Contact( #DeviceState.mySTATE[6] )
      Move(in := 100, out1 => #korak)
   END_RUNG
   // the same network as SCL:
   #trenutniKorak[45] := #korak = 45;
   IF (#korak = 45) AND #DeviceState.mySTATE[6] THEN #korak := 100; END_IF;
END_REGION

REGION Network 18: PRESTAVI HMI
   // Če je korak 100 -> prestavi HMI iz startupa
   // - če je HMI 17-> 0x11 = prestavi HMI
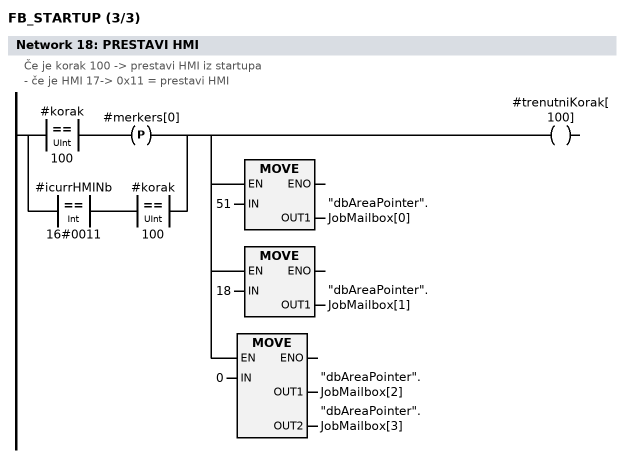
   RUNG wire#powerrail
      { S7_Templates := "SrcType := UInt" } EQ_Contact(in1 := #korak, in2 := 100)
      P_Trig( #merkers[0] )
      wire#w1
      Coil( #trenutniKorak[100] )
   END_RUNG
   RUNG wire#powerrail
      { S7_Templates := "SrcType := Int" } EQ_Contact(in1 := #icurrHMINb, in2 := 16#0011)
      { S7_Templates := "SrcType := UInt" } EQ_Contact(in1 := #korak, in2 := 100)
   END_RUNG wire#w1
   RUNG wire#w1
      Move(in := 51, out1 => "dbAreaPointer".JobMailbox[0])
   END_RUNG
   RUNG wire#w1
      Move(in := 18, out1 => "dbAreaPointer".JobMailbox[1])
   END_RUNG
   RUNG wire#w1
      Move(in := 0, out1 => "dbAreaPointer".JobMailbox[2], out2 => "dbAreaPointer".JobMailbox[3])
   END_RUNG
   // the same network as SCL:
   #_w1 := #korak = 100;
   #_w2 := #_w1 AND NOT #merkers[0];   // rising edge
   #merkers[0] := #_w1;
   #trenutniKorak[100] := #_w2 OR ((#icurrHMINb = 16#0011) AND (#korak = 100));
   IF #_w2 OR ((#icurrHMINb = 16#0011) AND (#korak = 100)) THEN
       "dbAreaPointer".JobMailbox[0] := 51;
       "dbAreaPointer".JobMailbox[1] := 18;
       "dbAreaPointer".JobMailbox[2] := 0;
       "dbAreaPointer".JobMailbox[3] := 0;
   END_IF;
END_REGION
END_FUNCTION_BLOCK

FUNCTION_BLOCK "FB_FESTO_SDE1"   // FB8, LAD
{ S7_Optimized_Access := 'TRUE' }
VERSION : 0.1
   VAR_INPUT
      iWord : UInt;
   END_VAR
   VAR_OUTPUT
      oPritisk : Real;
   END_VAR
   VAR CONSTANT
      "0BAR" : Real := 58620.0;
      "6BAR" : Real := 13997.0;
   END_VAR
BEGIN

REGION Network 2 (SCL)
   //4mA.....0bar
   //20mA....10bar
   //y := k*x + n

   #oPritisk := #"0BAR"/#"6BAR" * #iWord;
END_REGION
END_FUNCTION_BLOCK

FUNCTION_BLOCK "FB_ROČNO_VODENJE"   // FB11, LAD
{ S7_Optimized_Access := 'TRUE' }
VERSION : 0.1
   VAR_INPUT
      "TIPPEN_+" : Bool;
      "TIPPEN_-" : Bool;
      JeVRočnemNačinu : Bool;
      stCilindra : Int;
      iServoGo : Bool;
   END_VAR
   VAR_OUTPUT
      "Y1/1" : Bool;   // Zapora linearnega pogona / komada
      "Y2/1_1" : Bool;   // Vstavljanje nazaj
      "Y2/2_2" : Bool;   // Vstavljanje naprej
      "Y3/1" : Bool;   // CIlinder opridanje/zapiranje komada pri vstavljanju
      "Y1/2" : Bool;   // PobiranjePloščice
      "Y1/2_2" : Bool;   // NalaganjePloščice
      "Y1/4_1" : Bool;   // DvigElektrode
      "Y1/4_2" : Bool;   // SpustElektrode
      "Y2/3_1" : Bool;   // PoravnavaNaprej
      "Y2/3_2" : Bool;   // PoravnavaNazaj
      "Y3/1_1" : Bool;   // OdklepKonusa
      "Y3/3_1" : Bool;   // Odklep za vstavljanje izdelka
      "Y4/3_1" : Bool;   // Odklep izmeta izdelka
      Y5_3_1 : Bool;   // Izmet komada
      "Y6/3_1" : Bool;   // DrcaSlabi
      "Y6/3_2" : Bool;   // DrcaDobri
   END_VAR
   VAR_IN_OUT
      ServoGoVrtljivaMiza : Bool;
      ServoGoELektrodaZgoraj : Bool;
      ServoGoRezanjePodajajnje : Bool;
   END_VAR
   VAR
      IEC_Timer_0_Instance : TON_TIME;
      IEC_Timer_0_Instance_1 : TON_TIME;
      merkerji : Array[0..4] of Bool;
   END_VAR
   VAR_TEMP   // added for the SCL form of the ladder/FBD networks
      _w1 : Bool;
      _w2 : Bool;
      _w3 : Bool;
   END_VAR
BEGIN

REGION Network 1: ODKLEP/ZAKLEP LINISKEGA VIBRATORJA - 1y1
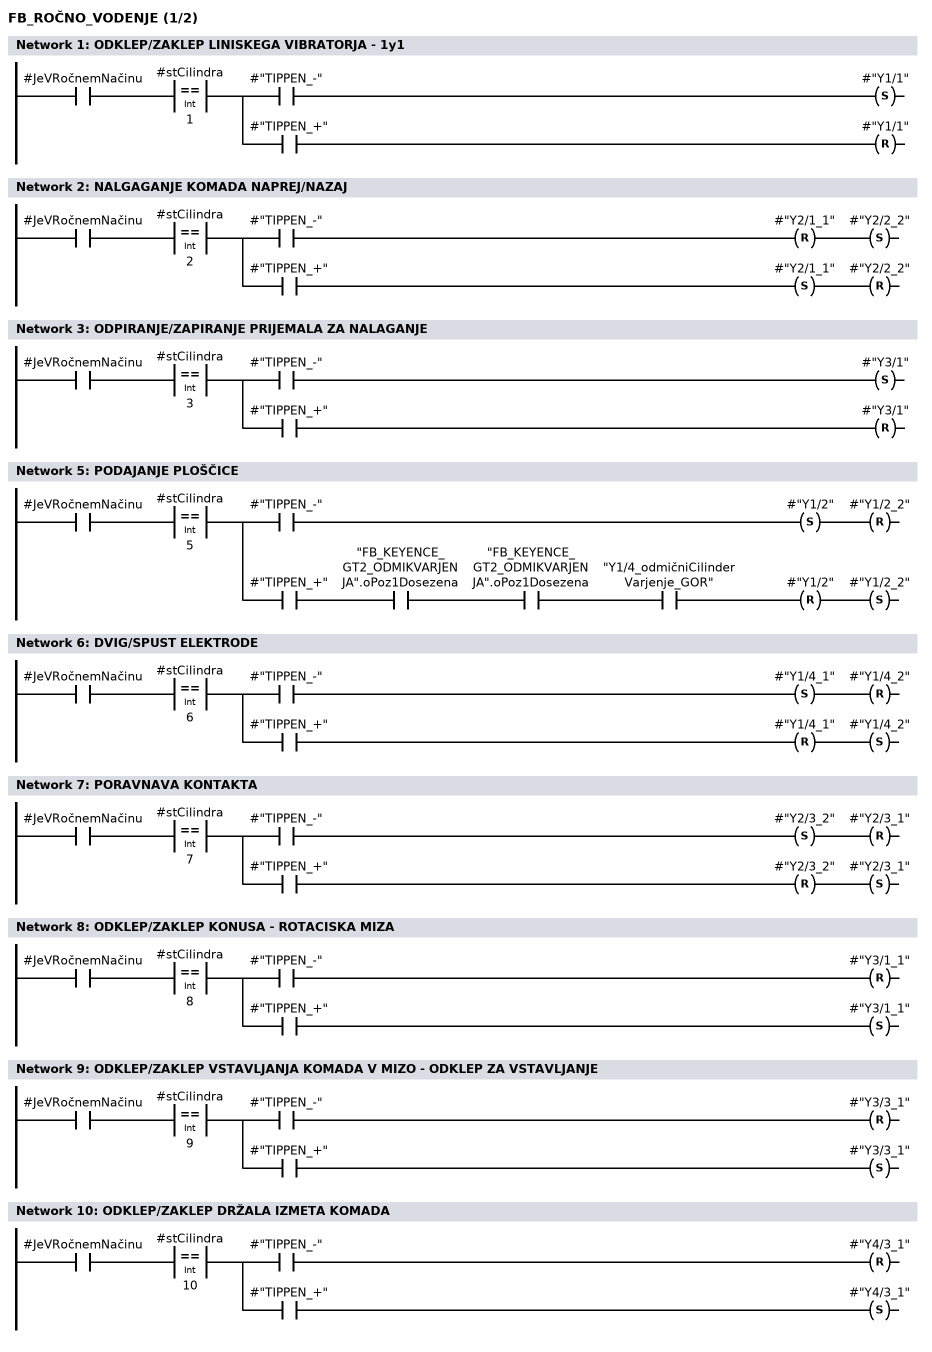
   RUNG wire#powerrail
      Contact( #JeVRočnemNačinu )
      { S7_Templates := "SrcType := Int" } EQ_Contact(in1 := #stCilindra, in2 := 1)
      wire#w1
      Contact( #"TIPPEN_-" )
      S_Coil( #"Y1/1" )
   END_RUNG
   RUNG wire#w1
      Contact( #"TIPPEN_+" )
      R_Coil( #"Y1/1" )
   END_RUNG
   // the same network as SCL:
   #_w1 := #JeVRočnemNačinu AND (#stCilindra = 1);
   IF #_w1 AND #"TIPPEN_-" THEN #"Y1/1" := TRUE; END_IF;
   IF #_w1 AND #"TIPPEN_+" THEN #"Y1/1" := FALSE; END_IF;
END_REGION

REGION Network 2: NALGAGANJE KOMADA NAPREJ/NAZAJ
   RUNG wire#powerrail
      Contact( #JeVRočnemNačinu )
      { S7_Templates := "SrcType := Int" } EQ_Contact(in1 := #stCilindra, in2 := 2)
      wire#w1
      Contact( #"TIPPEN_-" )
      R_Coil( #"Y2/1_1" )
      S_Coil( #"Y2/2_2" )
   END_RUNG
   RUNG wire#w1
      Contact( #"TIPPEN_+" )
      S_Coil( #"Y2/1_1" )
      R_Coil( #"Y2/2_2" )
   END_RUNG
   // the same network as SCL:
   #_w1 := #JeVRočnemNačinu AND (#stCilindra = 2);
   IF #_w1 AND #"TIPPEN_-" THEN
       #"Y2/1_1" := FALSE;
       #"Y2/2_2" := TRUE;
   END_IF;
   IF #_w1 AND #"TIPPEN_+" THEN
       #"Y2/1_1" := TRUE;
       #"Y2/2_2" := FALSE;
   END_IF;
END_REGION

REGION Network 3: ODPIRANJE/ZAPIRANJE PRIJEMALA ZA NALAGANJE
   RUNG wire#powerrail
      Contact( #JeVRočnemNačinu )
      { S7_Templates := "SrcType := Int" } EQ_Contact(in1 := #stCilindra, in2 := 3)
      wire#w1
      Contact( #"TIPPEN_-" )
      S_Coil( #"Y3/1" )
   END_RUNG
   RUNG wire#w1
      Contact( #"TIPPEN_+" )
      R_Coil( #"Y3/1" )
   END_RUNG
   // the same network as SCL:
   #_w1 := #JeVRočnemNačinu AND (#stCilindra = 3);
   IF #_w1 AND #"TIPPEN_-" THEN #"Y3/1" := TRUE; END_IF;
   IF #_w1 AND #"TIPPEN_+" THEN #"Y3/1" := FALSE; END_IF;
END_REGION
